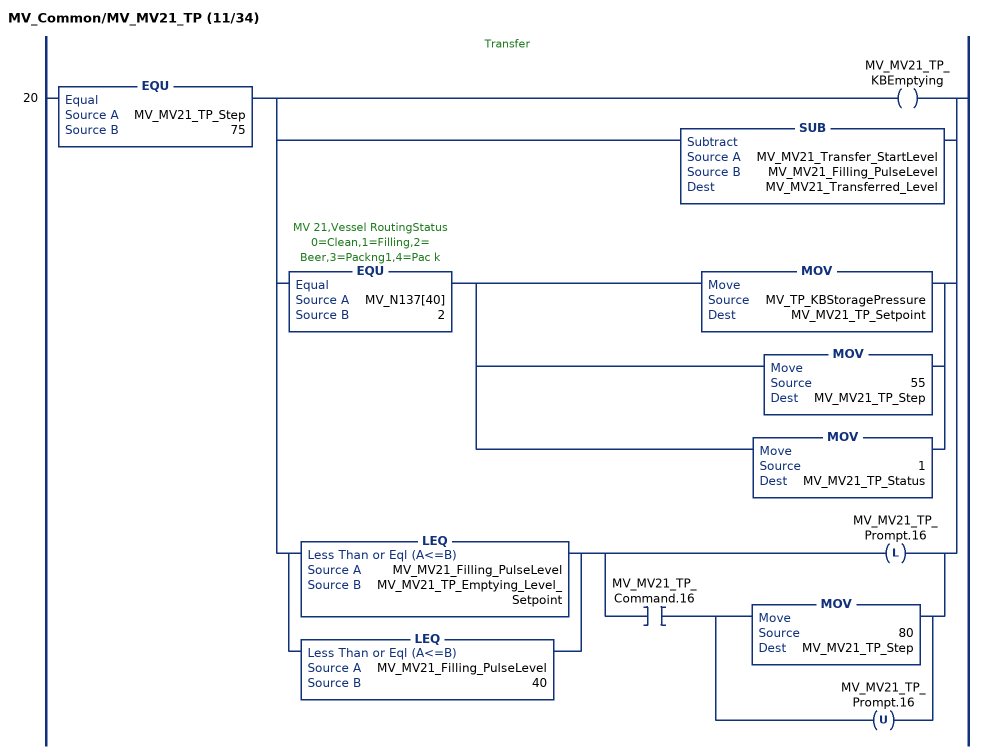
   // Transfer
   20: EQU(MV_MV21_TP_Step,75)[OTE(MV_MV21_TP_KBEmptying) ,SUB(MV_MV21_Transfer_StartLevel,MV_MV21_Filling_PulseLevel,MV_MV21_Transferred_Level) ,EQU(MV_N137[40],2) [MOV(MV_TP_KBStoragePressure,MV_MV21_TP_Setpoint) ,MOV(55,MV_MV21_TP_Step) ,MOV(1,MV_MV21_TP_Status) ] ,[LEQ(MV_MV21_Filling_PulseLevel,MV_MV21_TP_Emptying_Level_Setpoint) ,LEQ(MV_MV21_Filling_PulseLevel,40) ] [OTL(MV_MV21_TP_Prompt.16) ,XIC(MV_MV21_TP_Command.16) [MOV(80,MV_MV21_TP_Step) ,OTU(MV_MV21_TP_Prompt.16) ] ] ];
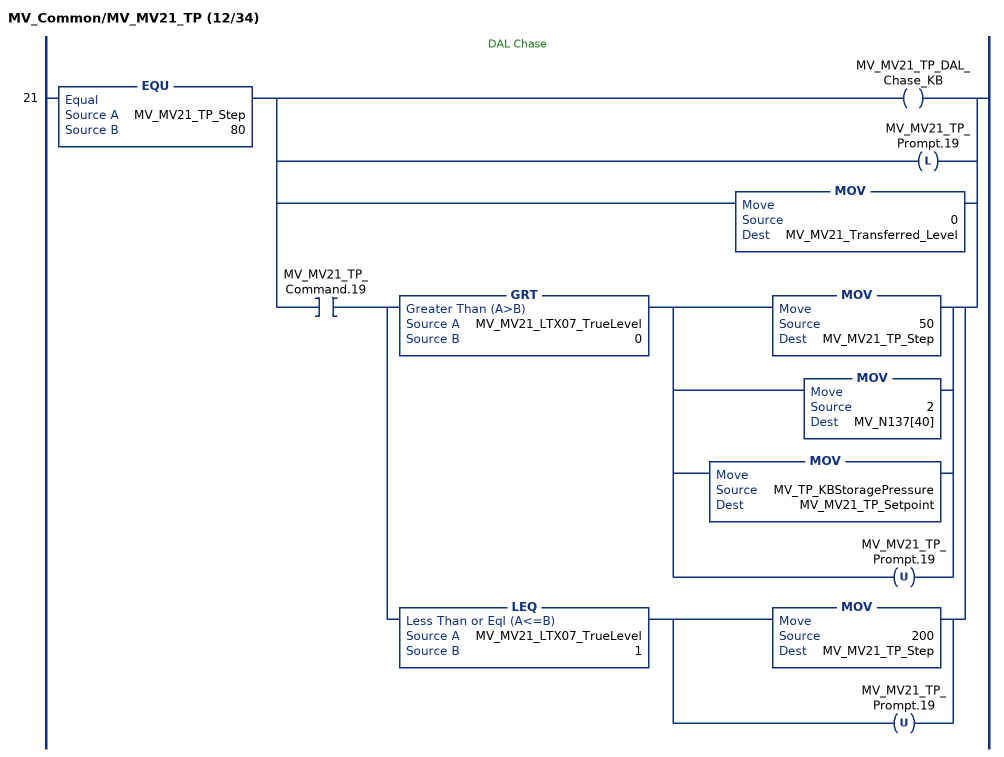
   // DAL Chase
   21: EQU(MV_MV21_TP_Step,80)[OTE(MV_MV21_TP_DAL_Chase_KB) ,OTL(MV_MV21_TP_Prompt.19) ,MOV(0,MV_MV21_Transferred_Level) ,XIC(MV_MV21_TP_Command.19) [GRT(MV_MV21_LTX07_TrueLevel,0) [MOV(50,MV_MV21_TP_Step) ,MOV(2,MV_N137[40]) ,MOV(MV_TP_KBStoragePressure,MV_MV21_TP_Setpoint) ,OTU(MV_MV21_TP_Prompt.19) ] ,LEQ(MV_MV21_LTX07_TrueLevel,1) [MOV(200,MV_MV21_TP_Step) ,OTU(MV_MV21_TP_Prompt.19) ] ] ];
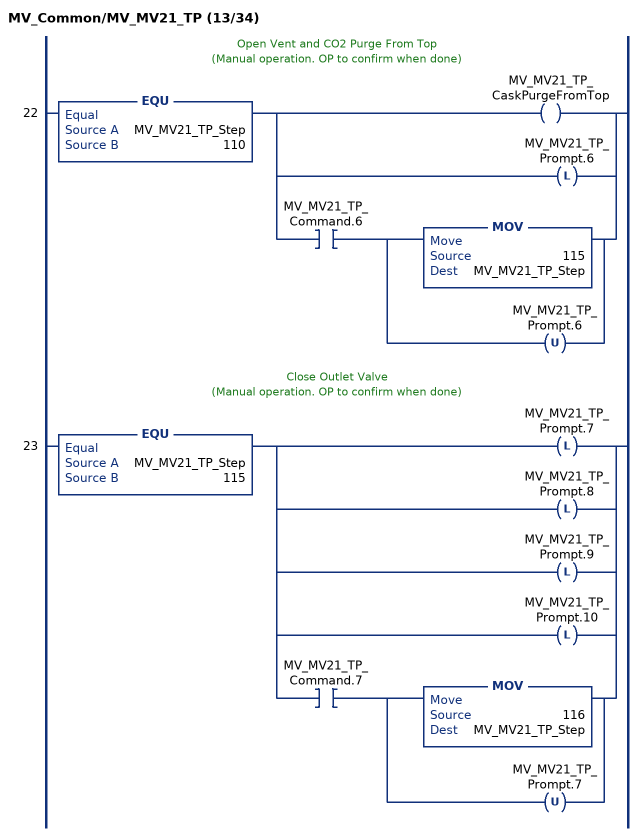
   // Open Vent and CO2 Purge From Top
   // (Manual operation. OP to confirm when done)
   22: EQU(MV_MV21_TP_Step,110)[OTE(MV_MV21_TP_CaskPurgeFromTop) ,OTL(MV_MV21_TP_Prompt.6) ,XIC(MV_MV21_TP_Command.6) [MOV(115,MV_MV21_TP_Step) ,OTU(MV_MV21_TP_Prompt.6) ] ];
   // Close Outlet Valve
   // (Manual operation. OP to confirm when done)
   23: EQU(MV_MV21_TP_Step,115)[OTL(MV_MV21_TP_Prompt.7) ,OTL(MV_MV21_TP_Prompt.8) ,OTL(MV_MV21_TP_Prompt.9) ,OTL(MV_MV21_TP_Prompt.10) ,XIC(MV_MV21_TP_Command.7) [MOV(116,MV_MV21_TP_Step) ,OTU(MV_MV21_TP_Prompt.7) ] ];
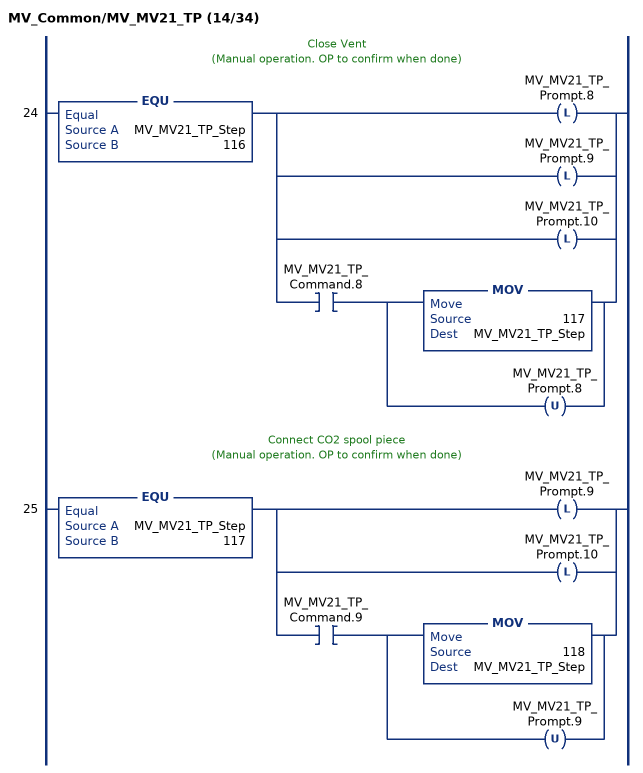
   // Close Vent
   // (Manual operation. OP to confirm when done)
   24: EQU(MV_MV21_TP_Step,116)[OTL(MV_MV21_TP_Prompt.8) ,OTL(MV_MV21_TP_Prompt.9) ,OTL(MV_MV21_TP_Prompt.10) ,XIC(MV_MV21_TP_Command.8) [MOV(117,MV_MV21_TP_Step) ,OTU(MV_MV21_TP_Prompt.8) ] ];
   // Connect CO2 spool piece
   // (Manual operation. OP to confirm when done)
   25: EQU(MV_MV21_TP_Step,117)[OTL(MV_MV21_TP_Prompt.9) ,OTL(MV_MV21_TP_Prompt.10) ,XIC(MV_MV21_TP_Command.9) [MOV(118,MV_MV21_TP_Step) ,OTU(MV_MV21_TP_Prompt.9) ] ];
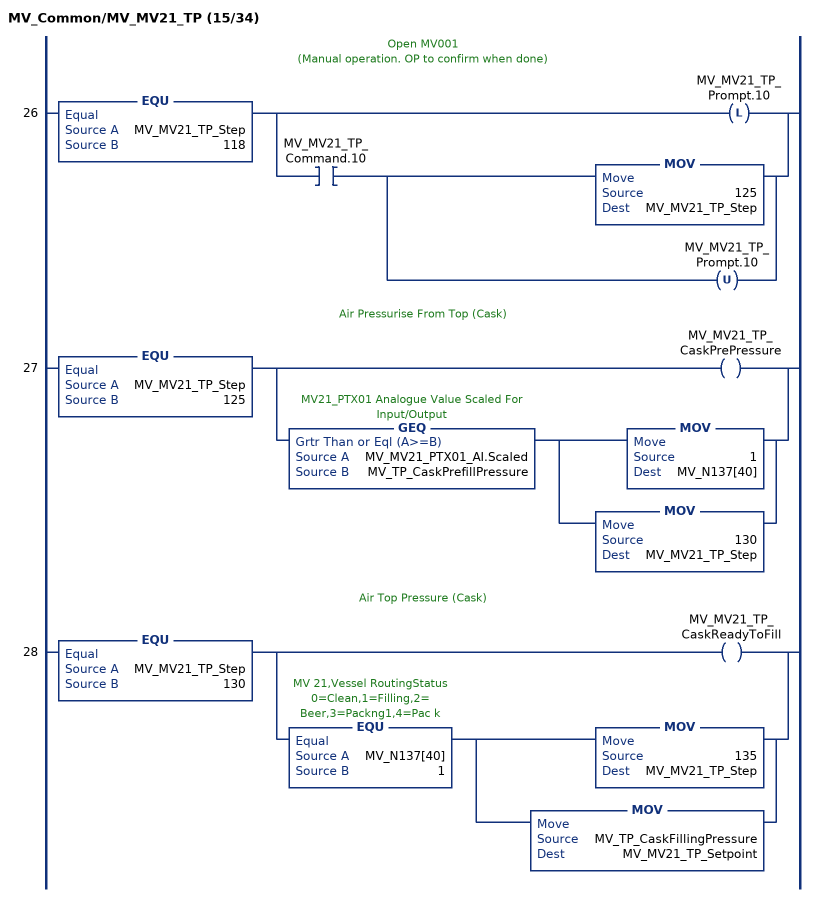
   // Open MV001
   // (Manual operation. OP to confirm when done)
   26: EQU(MV_MV21_TP_Step,118)[OTL(MV_MV21_TP_Prompt.10) ,XIC(MV_MV21_TP_Command.10) [MOV(125,MV_MV21_TP_Step) ,OTU(MV_MV21_TP_Prompt.10) ] ];
   // Air Pressurise From Top (Cask)
   27: EQU(MV_MV21_TP_Step,125)[OTE(MV_MV21_TP_CaskPrePressure) ,GEQ(MV_MV21_PTX01_AI.Scaled,MV_TP_CaskPrefillPressure) [MOV(1,MV_N137[40]) ,MOV(130,MV_MV21_TP_Step) ] ];
   // Air Top Pressure (Cask)
   28: EQU(MV_MV21_TP_Step,130)[OTE(MV_MV21_TP_CaskReadyToFill) ,EQU(MV_N137[40],1) [MOV(135,MV_MV21_TP_Step) ,MOV(MV_TP_CaskFillingPressure,MV_MV21_TP_Setpoint) ] ];
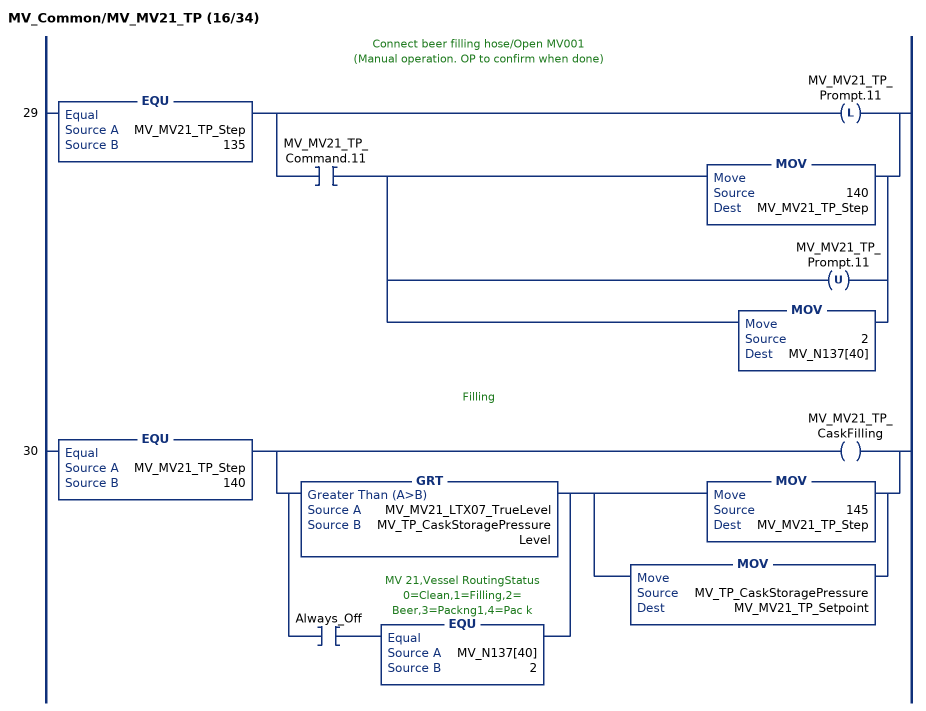
   // Connect beer filling hose/Open MV001
   // (Manual operation. OP to confirm when done)
   29: EQU(MV_MV21_TP_Step,135)[OTL(MV_MV21_TP_Prompt.11) ,XIC(MV_MV21_TP_Command.11) [MOV(140,MV_MV21_TP_Step) ,OTU(MV_MV21_TP_Prompt.11) ,MOV(2,MV_N137[40]) ] ];
   // Filling
   30: EQU(MV_MV21_TP_Step,140)[OTE(MV_MV21_TP_CaskFilling) ,[GRT(MV_MV21_LTX07_TrueLevel,MV_TP_CaskStoragePressureLevel) ,XIC(Always_Off) EQU(MV_N137[40],2) ] [MOV(145,MV_MV21_TP_Step) ,MOV(MV_TP_CaskStoragePressure,MV_MV21_TP_Setpoint) ] ];
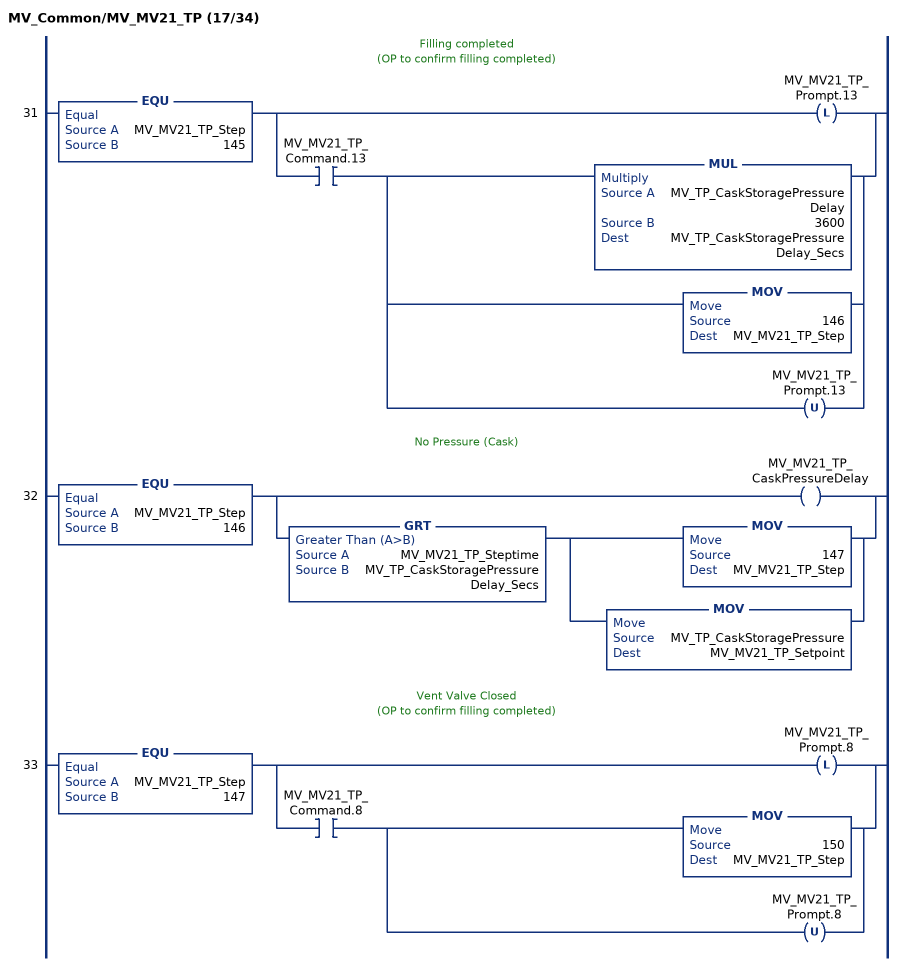
   // Filling completed
   // (OP to confirm filling completed)
   31: EQU(MV_MV21_TP_Step,145)[OTL(MV_MV21_TP_Prompt.13) ,XIC(MV_MV21_TP_Command.13) [MUL(MV_TP_CaskStoragePressureDelay,3600,MV_TP_CaskStoragePressureDelay_Secs) ,MOV(146,MV_MV21_TP_Step) ,OTU(MV_MV21_TP_Prompt.13) ] ];
   // No Pressure (Cask)
   32: EQU(MV_MV21_TP_Step,146)[OTE(MV_MV21_TP_CaskPressureDelay) ,GRT(MV_MV21_TP_Steptime,MV_TP_CaskStoragePressureDelay_Secs) [MOV(147,MV_MV21_TP_Step) ,MOV(MV_TP_CaskStoragePressure,MV_MV21_TP_Setpoint) ] ];
   // Vent Valve Closed
   // (OP to confirm filling completed)
   33: EQU(MV_MV21_TP_Step,147)[OTL(MV_MV21_TP_Prompt.8) ,XIC(MV_MV21_TP_Command.8) [MOV(150,MV_MV21_TP_Step) ,OTU(MV_MV21_TP_Prompt.8) ] ];
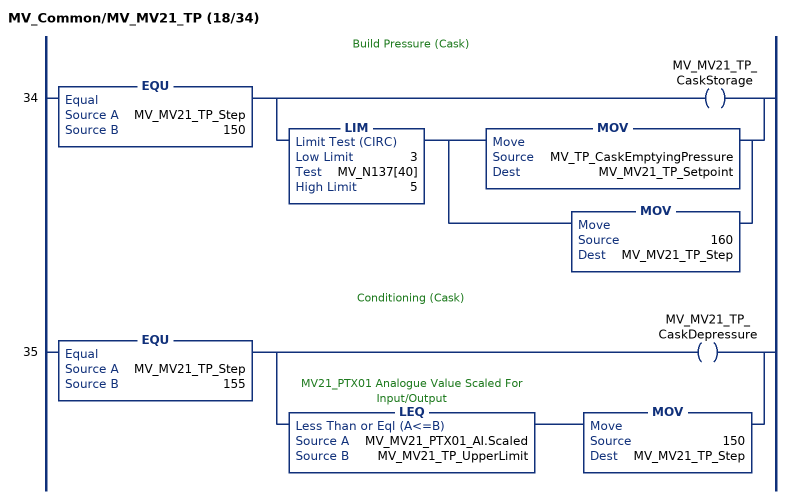
   // Build Pressure (Cask)
   34: EQU(MV_MV21_TP_Step,150)[OTE(MV_MV21_TP_CaskStorage) ,LIM(3,MV_N137[40],5) [MOV(MV_TP_CaskEmptyingPressure,MV_MV21_TP_Setpoint) ,MOV(160,MV_MV21_TP_Step) ] ];
   // Conditioning (Cask)
   35: EQU(MV_MV21_TP_Step,155)[OTE(MV_MV21_TP_CaskDepressure) ,LEQ(MV_MV21_PTX01_AI.Scaled,MV_MV21_TP_UpperLimit) MOV(150,MV_MV21_TP_Step) ];
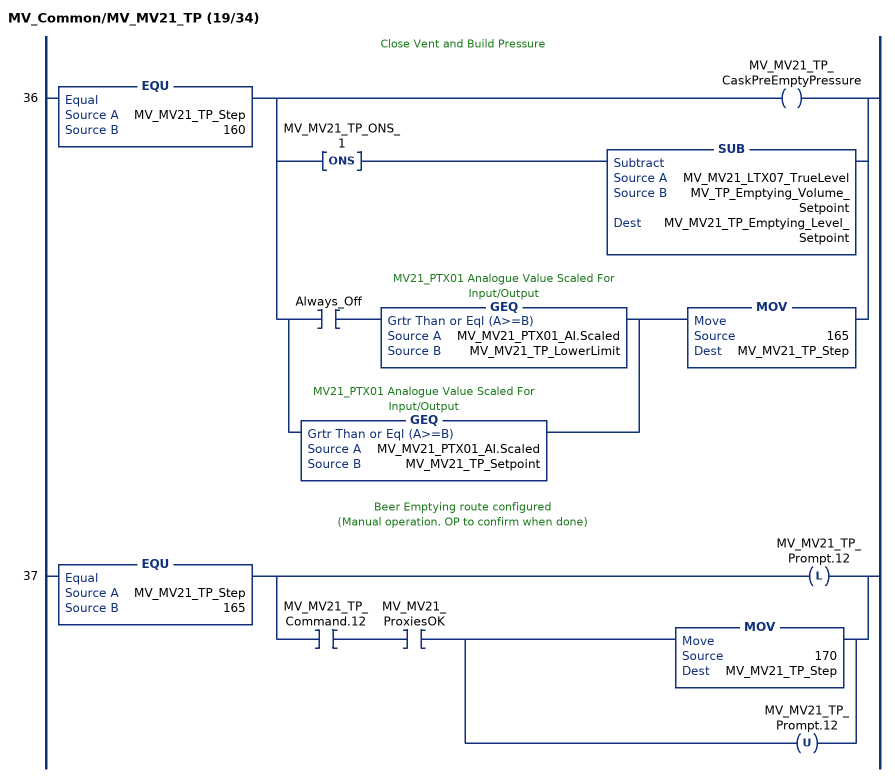
   // Close Vent and Build Pressure
   36: EQU(MV_MV21_TP_Step,160)[OTE(MV_MV21_TP_CaskPreEmptyPressure) ,ONS(MV_MV21_TP_ONS_1) SUB(MV_MV21_LTX07_TrueLevel,MV_TP_Emptying_Volume_Setpoint,MV_MV21_TP_Emptying_Level_Setpoint) ,[XIC(Always_Off) GEQ(MV_MV21_PTX01_AI.Scaled,MV_MV21_TP_LowerLimit) ,GEQ(MV_MV21_PTX01_AI.Scaled,MV_MV21_TP_Setpoint) ] MOV(165,MV_MV21_TP_Step) ];
   // Beer Emptying route configured
   // (Manual operation. OP to confirm when done)
   37: EQU(MV_MV21_TP_Step,165)[OTL(MV_MV21_TP_Prompt.12) ,XIC(MV_MV21_TP_Command.12) XIC(MV_MV21_ProxiesOK) [MOV(170,MV_MV21_TP_Step) ,OTU(MV_MV21_TP_Prompt.12) ] ];
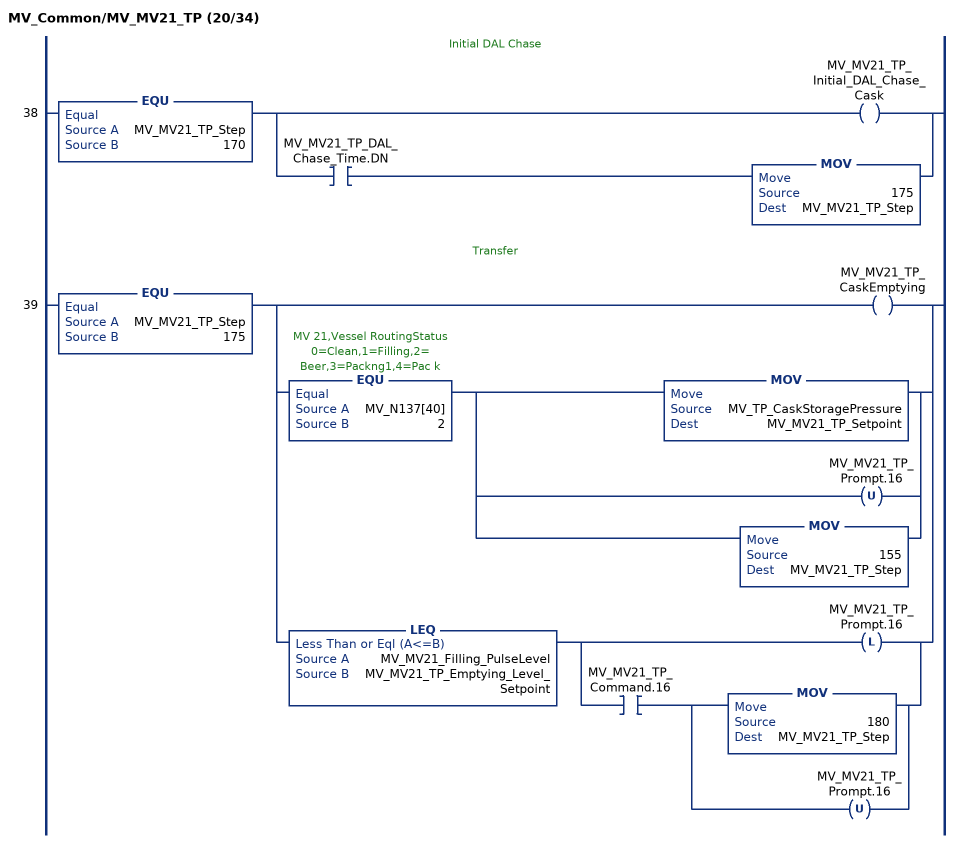
   // Initial DAL Chase
   38: EQU(MV_MV21_TP_Step,170)[OTE(MV_MV21_TP_Initial_DAL_Chase_Cask) ,XIC(MV_MV21_TP_DAL_Chase_Time.DN) MOV(175,MV_MV21_TP_Step) ];
   // Transfer
   39: EQU(MV_MV21_TP_Step,175)[OTE(MV_MV21_TP_CaskEmptying) ,EQU(MV_N137[40],2) [MOV(MV_TP_CaskStoragePressure,MV_MV21_TP_Setpoint) ,OTU(MV_MV21_TP_Prompt.16) ,MOV(155,MV_MV21_TP_Step) ] ,LEQ(MV_MV21_Filling_PulseLevel,MV_MV21_TP_Emptying_Level_Setpoint) [OTL(MV_MV21_TP_Prompt.16) ,XIC(MV_MV21_TP_Command.16) [MOV(180,MV_MV21_TP_Step) ,OTU(MV_MV21_TP_Prompt.16) ] ] ];
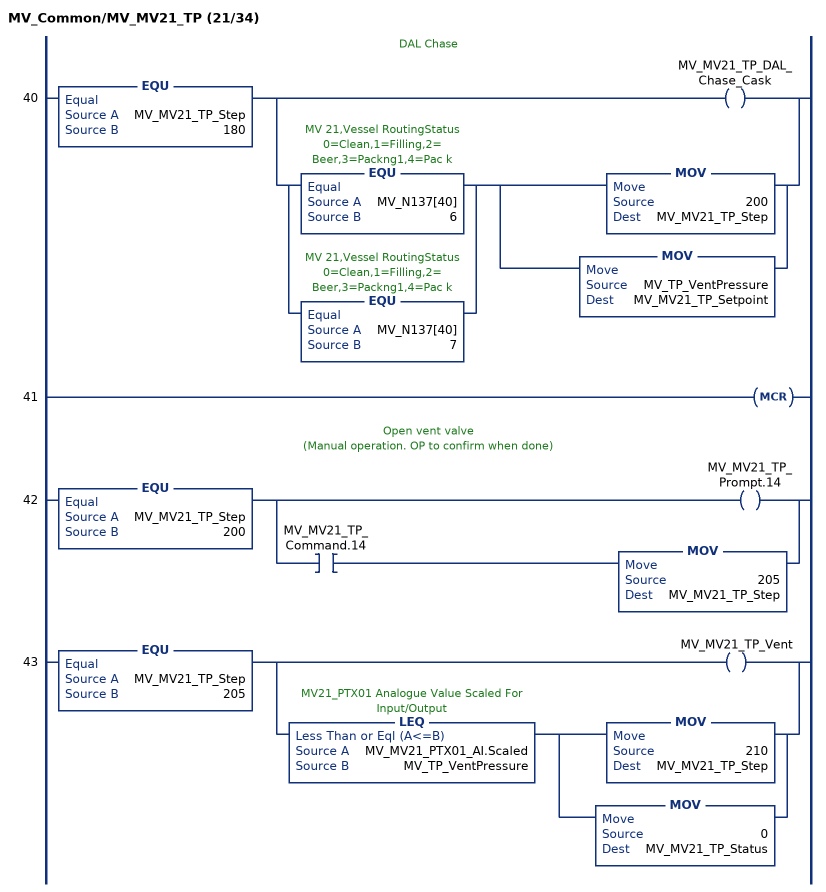
   // DAL Chase
   40: EQU(MV_MV21_TP_Step,180)[OTE(MV_MV21_TP_DAL_Chase_Cask) ,[EQU(MV_N137[40],6) ,EQU(MV_N137[40],7) ] [MOV(200,MV_MV21_TP_Step) ,MOV(MV_TP_VentPressure,MV_MV21_TP_Setpoint) ] ];
   41: MCR();
   // Open vent valve
   // (Manual operation. OP to confirm when done)
   42: EQU(MV_MV21_TP_Step,200)[OTE(MV_MV21_TP_Prompt.14) ,XIC(MV_MV21_TP_Command.14) MOV(205,MV_MV21_TP_Step) ];
   43: EQU(MV_MV21_TP_Step,205)[OTE(MV_MV21_TP_Vent) ,LEQ(MV_MV21_PTX01_AI.Scaled,MV_TP_VentPressure) [MOV(210,MV_MV21_TP_Step) ,MOV(0,MV_MV21_TP_Status) ] ];
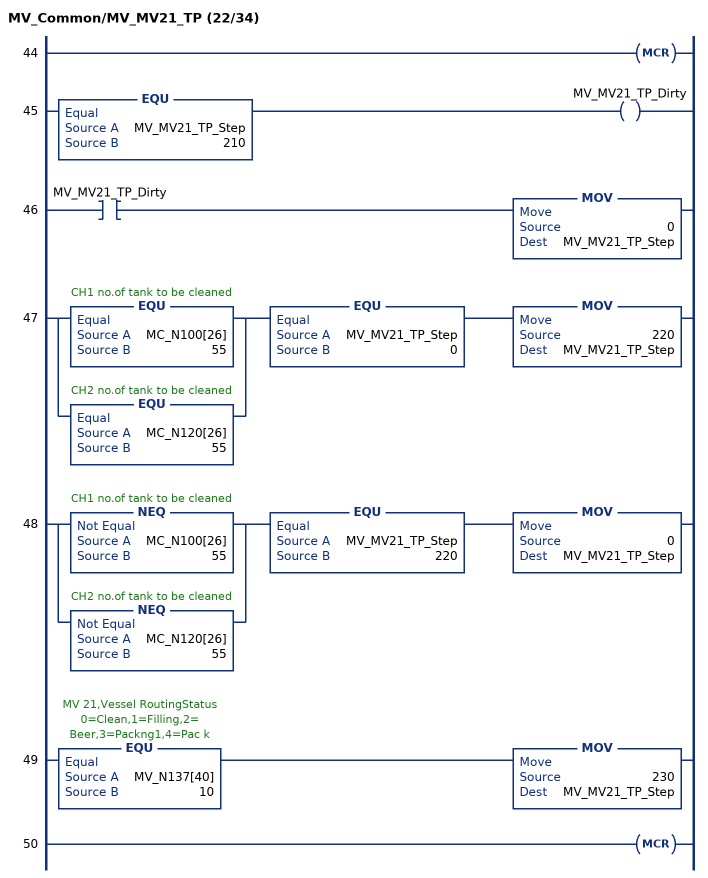
   44: MCR();
   45: EQU(MV_MV21_TP_Step,210)OTE(MV_MV21_TP_Dirty);
   46: XIC(MV_MV21_TP_Dirty)MOV(0,MV_MV21_TP_Step);
   47: [EQU(MC_N100[26],55) ,EQU(MC_N120[26],55) ]EQU(MV_MV21_TP_Step,0)MOV(220,MV_MV21_TP_Step);
   48: [NEQ(MC_N100[26],55) ,NEQ(MC_N120[26],55) ]EQU(MV_MV21_TP_Step,220)MOV(0,MV_MV21_TP_Step);
   49: EQU(MV_N137[40],10)MOV(230,MV_MV21_TP_Step);
   50: MCR();
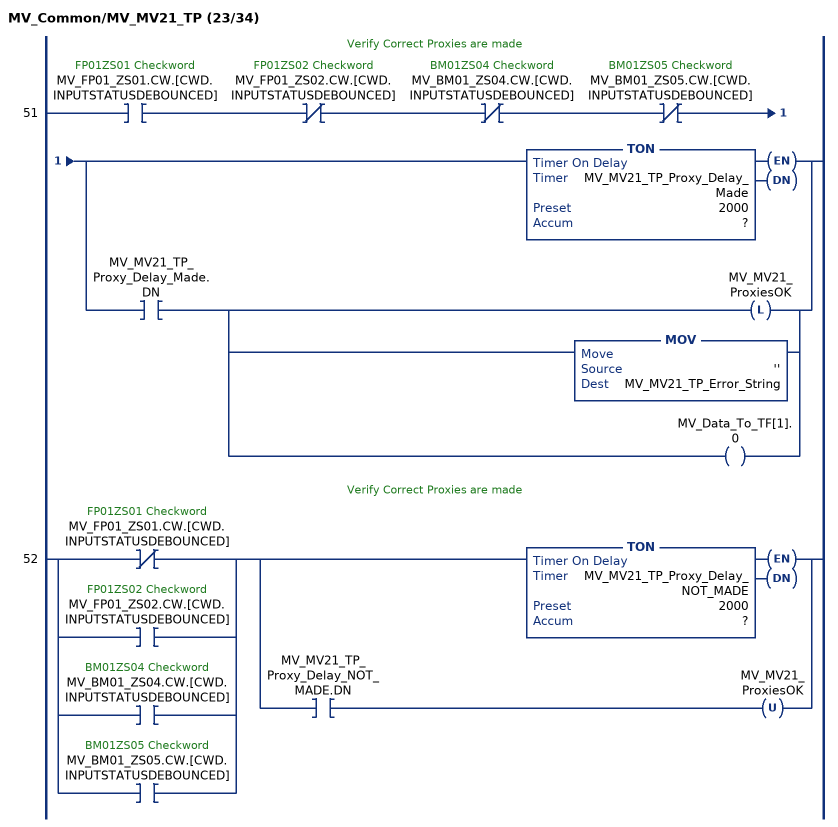
   // Verify Correct Proxies are made
   51: XIC(MV_FP01_ZS01.CW.[CWD.INPUTSTATUSDEBOUNCED])XIO(MV_FP01_ZS02.CW.[CWD.INPUTSTATUSDEBOUNCED])XIO(MV_BM01_ZS04.CW.[CWD.INPUTSTATUSDEBOUNCED])XIO(MV_BM01_ZS05.CW.[CWD.INPUTSTATUSDEBOUNCED])[TON(MV_MV21_TP_Proxy_Delay_Made,?,?) ,XIC(MV_MV21_TP_Proxy_Delay_Made.DN) [OTL(MV_MV21_ProxiesOK) ,MOV('',MV_MV21_TP_Error_String) ,OTE(MV_Data_To_TF[1].0) ] ];
   // Verify Correct Proxies are made
   52: [XIO(MV_FP01_ZS01.CW.[CWD.INPUTSTATUSDEBOUNCED]) ,XIC(MV_FP01_ZS02.CW.[CWD.INPUTSTATUSDEBOUNCED]) ,XIC(MV_BM01_ZS04.CW.[CWD.INPUTSTATUSDEBOUNCED]) ,XIC(MV_BM01_ZS05.CW.[CWD.INPUTSTATUSDEBOUNCED]) ][TON(MV_MV21_TP_Proxy_Delay_NOT_MADE,?,?) ,XIC(MV_MV21_TP_Proxy_Delay_NOT_MADE.DN) OTU(MV_MV21_ProxiesOK) ];
